   "Carrier_66_Motion_On_Fault" AT %Q3676.5 : Bool;
   "Carrier_66_Motion_Off_Fault" AT %Q3676.6 : Bool;
   "Carrier_66_Carrier_Spacing_Fault" AT %Q3676.7 : Bool;
   "Carrier_67_Carrier_In_Zone" AT %QW3700 : Word;
   "Carrier_67_Carrier_Number_Echo" AT %QW3702 : Word;
   "Carrier_67_Carrier_Position_Echo" AT %QD3704 : DWord;
   "Carrier_67_Next_Carrier_Number" AT %QW3708 : Word;
   "Carrier_67_Next_Stop_Position" AT %QD3710 : DWord;
   "Carrier_67_Drive_Command_Speed" AT %QW3714 : Word;
   "Carrier_67_Duplicate_Carrier_Number" AT %QW3716 : Word;
   "Carrier_67_First_Duplicate_Carrier_Position" AT %QD3718 : DWord;
   "Carrier_67_Second_Duplicate_Carrier_Position" AT %QD3722 : DWord;
   "Carrier_67_CommandWord" AT %QW3726 : Word;
   "Carrier_67_Heartbeat" AT %Q3726.0 : Bool;
   "Carrier_67_Drive_Forward_Command" AT %Q3726.1 : Bool;
   "Carrier_67_Fault_Reset" AT %Q3726.2 : Bool;
   "Carrier_67_At_Command_Position" AT %Q3726.3 : Bool;
   "Carrier_67_Duplicate_Carrier_Fault" AT %Q3726.4 : Bool;
   "Carrier_67_Motion_On_Fault" AT %Q3726.5 : Bool;
   "Carrier_67_Motion_Off_Fault" AT %Q3726.6 : Bool;
   "Carrier_67_Carrier_Spacing_Fault" AT %Q3726.7 : Bool;
   "Carrier_68_Carrier_In_Zone" AT %QW3750 : Word;
   "Carrier_68_Carrier_Number_Echo" AT %QW3752 : Word;
   "Carrier_68_Carrier_Position_Echo" AT %QD3754 : DWord;
   "Carrier_68_Next_Carrier_Number" AT %QW3758 : Word;
   "Carrier_68_Next_Stop_Position" AT %QD3760 : DWord;
   "Carrier_68_Drive_Command_Speed" AT %QW3764 : Word;
   "Carrier_68_Duplicate_Carrier_Number" AT %QW3766 : Word;
   "Carrier_68_First_Duplicate_Carrier_Position" AT %QD3768 : DWord;
   "Carrier_68_Second_Duplicate_Carrier_Position" AT %QD3772 : DWord;
   "Carrier_68_CommandWord" AT %QW3776 : Word;
   "Carrier_68_Heartbeat" AT %Q3776.0 : Bool;
   "Carrier_68_Drive_Forward_Command" AT %Q3776.1 : Bool;
   "Carrier_68_Fault_Reset" AT %Q3776.2 : Bool;
   "Carrier_68_At_Command_Position" AT %Q3776.3 : Bool;
   "Carrier_68_Duplicate_Carrier_Fault" AT %Q3776.4 : Bool;
   "Carrier_68_Motion_On_Fault" AT %Q3776.5 : Bool;
   "Carrier_68_Motion_Off_Fault" AT %Q3776.6 : Bool;
   "Carrier_68_Carrier_Spacing_Fault" AT %Q3776.7 : Bool;
   "Carrier_69_Carrier_In_Zone" AT %QW3800 : Word;
   "Carrier_69_Carrier_Number_Echo" AT %QW3802 : Word;
   "Carrier_69_Carrier_Position_Echo" AT %QD3804 : DWord;
   "Carrier_69_Next_Carrier_Number" AT %QW3808 : Word;
   "Carrier_69_Next_Stop_Position" AT %QD3810 : DWord;
   "Carrier_69_Drive_Command_Speed" AT %QW3814 : Word;
   "Carrier_69_Duplicate_Carrier_Number" AT %QW3816 : Word;
   "Carrier_69_First_Duplicate_Carrier_Position" AT %QD3818 : DWord;
   "Carrier_69_Second_Duplicate_Carrier_Position" AT %QD3822 : DWord;
   "Carrier_69_CommandWord" AT %QW3826 : Word;
   "Carrier_69_Heartbeat" AT %Q3826.0 : Bool;
   "Carrier_69_Drive_Forward_Command" AT %Q3826.1 : Bool;
   "Carrier_69_Fault_Reset" AT %Q3826.2 : Bool;
   "Carrier_69_At_Command_Position" AT %Q3826.3 : Bool;
   "Carrier_69_Duplicate_Carrier_Fault" AT %Q3826.4 : Bool;
   "Carrier_69_Motion_On_Fault" AT %Q3826.5 : Bool;
   "Carrier_69_Motion_Off_Fault" AT %Q3826.6 : Bool;
   "Carrier_69_Carrier_Spacing_Fault" AT %Q3826.7 : Bool;
   "Carrier_70_Carrier_In_Zone" AT %QW3850 : Word;
   "Carrier_70_Carrier_Number_Echo" AT %QW3852 : Word;
   "Carrier_70_Carrier_Position_Echo" AT %QD3854 : DWord;
   "Carrier_70_Next_Carrier_Number" AT %QW3858 : Word;
   "Carrier_70_Next_Stop_Position" AT %QD3860 : DWord;
   "Carrier_70_Drive_Command_Speed" AT %QW3864 : Word;
   "Carrier_70_Duplicate_Carrier_Number" AT %QW3866 : Word;
   "Carrier_70_First_Duplicate_Carrier_Position" AT %QD3868 : DWord;
   "Carrier_70_Second_Duplicate_Carrier_Position" AT %QD3872 : DWord;
   "Carrier_70_CommandWord" AT %QW3876 : Word;
   "Carrier_70_Heartbeat" AT %Q3876.0 : Bool;
   "Carrier_70_Drive_Forward_Command" AT %Q3876.1 : Bool;
   "Carrier_70_Fault_Reset" AT %Q3876.2 : Bool;
   "Carrier_70_At_Command_Position" AT %Q3876.3 : Bool;
   "Carrier_70_Duplicate_Carrier_Fault" AT %Q3876.4 : Bool;
   "Carrier_70_Motion_On_Fault" AT %Q3876.5 : Bool;
   "Carrier_70_Motion_Off_Fault" AT %Q3876.6 : Bool;
   "Carrier_70_Carrier_Spacing_Fault" AT %Q3876.7 : Bool;
   "Carrier_71_Carrier_In_Zone" AT %QW3900 : Word;
   "Carrier_71_Carrier_Number_Echo" AT %QW3902 : Word;
   "Carrier_71_Carrier_Position_Echo" AT %QD3904 : DWord;
   "Carrier_71_Next_Carrier_Number" AT %QW3908 : Word;
   "Carrier_71_Next_Stop_Position" AT %QD3910 : DWord;
   "Carrier_71_Drive_Command_Speed" AT %QW3914 : Word;
   "Carrier_71_Duplicate_Carrier_Number" AT %QW3916 : Word;
   "Carrier_71_First_Duplicate_Carrier_Position" AT %QD3918 : DWord;
   "Carrier_71_Second_Duplicate_Carrier_Position" AT %QD3922 : DWord;
   "Carrier_71_CommandWord" AT %QW3926 : Word;
   "Carrier_71_Heartbeat" AT %Q3926.0 : Bool;
   "Carrier_71_Drive_Forward_Command" AT %Q3926.1 : Bool;
   "Carrier_71_Fault_Reset" AT %Q3926.2 : Bool;
   "Carrier_71_At_Command_Position" AT %Q3926.3 : Bool;
   "Carrier_71_Duplicate_Carrier_Fault" AT %Q3926.4 : Bool;
   "Carrier_71_Motion_On_Fault" AT %Q3926.5 : Bool;
   "Carrier_71_Motion_Off_Fault" AT %Q3926.6 : Bool;
   "Carrier_71_Carrier_Spacing_Fault" AT %Q3926.7 : Bool;
   "Carrier_72_Carrier_In_Zone" AT %QW3950 : Word;
   "Carrier_72_Carrier_Number_Echo" AT %QW3952 : Word;
   "Carrier_72_Carrier_Position_Echo" AT %QD3954 : DWord;
   "Carrier_72_Next_Carrier_Number" AT %QW3958 : Word;
   "Carrier_72_Next_Stop_Position" AT %QD3960 : DWord;
   "Carrier_72_Drive_Command_Speed" AT %QW3964 : Word;
   "Carrier_72_Duplicate_Carrier_Number" AT %QW3966 : Word;
   "Carrier_72_First_Duplicate_Carrier_Position" AT %QD3968 : DWord;
   "Carrier_72_Second_Duplicate_Carrier_Position" AT %QD3972 : DWord;
   "Carrier_72_CommandWord" AT %QW3976 : Word;
   "Carrier_72_Heartbeat" AT %Q3976.0 : Bool;
   "Carrier_72_Drive_Forward_Command" AT %Q3976.1 : Bool;
   "Carrier_72_Fault_Reset" AT %Q3976.2 : Bool;
   "Carrier_72_At_Command_Position" AT %Q3976.3 : Bool;
   "Carrier_72_Duplicate_Carrier_Fault" AT %Q3976.4 : Bool;
   "Carrier_72_Motion_On_Fault" AT %Q3976.5 : Bool;
   "Carrier_72_Motion_Off_Fault" AT %Q3976.6 : Bool;
   "Carrier_72_Carrier_Spacing_Fault" AT %Q3976.7 : Bool;
   "Carrier_73_Carrier_In_Zone" AT %QW4000 : Word;
   "Carrier_73_Carrier_Number_Echo" AT %QW4002 : Word;
   "Carrier_73_Carrier_Position_Echo" AT %QD4004 : DWord;
   "Carrier_73_Next_Carrier_Number" AT %QW4008 : Word;
   "Carrier_73_Next_Stop_Position" AT %QD4010 : DWord;
   "Carrier_73_Drive_Command_Speed" AT %QW4014 : Word;
   "Carrier_73_Duplicate_Carrier_Number" AT %QW4016 : Word;
   "Carrier_73_First_Duplicate_Carrier_Position" AT %QD4018 : DWord;
   "Carrier_73_Second_Duplicate_Carrier_Position" AT %QD4022 : DWord;
   "Carrier_73_CommandWord" AT %QW4026 : Word;
   "Carrier_73_Heartbeat" AT %Q4026.0 : Bool;
   "Carrier_73_Drive_Forward_Command" AT %Q4026.1 : Bool;
   "Carrier_73_Fault_Reset" AT %Q4026.2 : Bool;
   "Carrier_73_At_Command_Position" AT %Q4026.3 : Bool;
   "Carrier_73_Duplicate_Carrier_Fault" AT %Q4026.4 : Bool;
   "Carrier_73_Motion_On_Fault" AT %Q4026.5 : Bool;
   "Carrier_73_Motion_Off_Fault" AT %Q4026.6 : Bool;
   "Carrier_73_Carrier_Spacing_Fault" AT %Q4026.7 : Bool;
   "Carrier_74_Carrier_In_Zone" AT %QW4050 : Word;
   "Carrier_74_Carrier_Number_Echo" AT %QW4052 : Word;
   "Carrier_74_Carrier_Position_Echo" AT %QD4054 : DWord;
   "Carrier_74_Next_Carrier_Number" AT %QW4058 : Word;
   "Carrier_74_Next_Stop_Position" AT %QD4060 : DWord;
   "Carrier_74_Drive_Command_Speed" AT %QW4064 : Word;
   "Carrier_74_Duplicate_Carrier_Number" AT %QW4066 : Word;
   "Carrier_74_First_Duplicate_Carrier_Position" AT %QD4068 : DWord;
   "Carrier_74_Second_Duplicate_Carrier_Position" AT %QD4072 : DWord;
   "Carrier_74_CommandWord" AT %QW4076 : Word;
   "Carrier_74_Heartbeat" AT %Q4076.0 : Bool;
   "Carrier_74_Drive_Forward_Command" AT %Q4076.1 : Bool;
   "Carrier_74_Fault_Reset" AT %Q4076.2 : Bool;
   "Carrier_74_At_Command_Position" AT %Q4076.3 : Bool;
   "Carrier_74_Duplicate_Carrier_Fault" AT %Q4076.4 : Bool;
   "Carrier_74_Motion_On_Fault" AT %Q4076.5 : Bool;
   "Carrier_74_Motion_Off_Fault" AT %Q4076.6 : Bool;
   "Carrier_74_Carrier_Spacing_Fault" AT %Q4076.7 : Bool;
   "Carrier_75_Carrier_In_Zone" AT %QW4100 : Word;
   "Carrier_75_Carrier_Number_Echo" AT %QW4102 : Word;
   "Carrier_75_Carrier_Position_Echo" AT %QD4104 : DWord;
   "Carrier_75_Next_Carrier_Number" AT %QW4108 : Word;
   "Carrier_75_Next_Stop_Position" AT %QD4110 : DWord;
   "Carrier_75_Drive_Command_Speed" AT %QW4114 : Word;
   "Carrier_75_Duplicate_Carrier_Number" AT %QW4116 : Word;
   "Carrier_75_First_Duplicate_Carrier_Position" AT %QD4118 : DWord;
   "Carrier_75_Second_Duplicate_Carrier_Position" AT %QD4122 : DWord;
   "Carrier_75_CommandWord" AT %QW4126 : Word;
   "Carrier_75_Heartbeat" AT %Q4126.0 : Bool;
   "Carrier_75_Drive_Forward_Command" AT %Q4126.1 : Bool;
   "Carrier_75_Fault_Reset" AT %Q4126.2 : Bool;
   "Carrier_75_At_Command_Position" AT %Q4126.3 : Bool;
   "Carrier_75_Duplicate_Carrier_Fault" AT %Q4126.4 : Bool;
   "Carrier_75_Motion_On_Fault" AT %Q4126.5 : Bool;
   "Carrier_75_Motion_Off_Fault" AT %Q4126.6 : Bool;
   "Carrier_75_Carrier_Spacing_Fault" AT %Q4126.7 : Bool;
   "Carrier_76_Carrier_In_Zone" AT %QW4150 : Word;
   "Carrier_76_Carrier_Number_Echo" AT %QW4152 : Word;
   "Carrier_76_Carrier_Position_Echo" AT %QD4154 : DWord;
   "Carrier_76_Next_Carrier_Number" AT %QW4158 : Word;
   "Carrier_76_Next_Stop_Position" AT %QD4160 : DWord;
   "Carrier_76_Drive_Command_Speed" AT %QW4164 : Word;
   "Carrier_76_Duplicate_Carrier_Number" AT %QW4166 : Word;
   "Carrier_76_First_Duplicate_Carrier_Position" AT %QD4168 : DWord;
   "Carrier_76_Second_Duplicate_Carrier_Position" AT %QD4172 : DWord;
   "Carrier_76_CommandWord" AT %QW4176 : Word;
   "Carrier_76_Heartbeat" AT %Q4176.0 : Bool;
   "Carrier_76_Drive_Forward_Command" AT %Q4176.1 : Bool;
   "Carrier_76_Fault_Reset" AT %Q4176.2 : Bool;
   "Carrier_76_At_Command_Position" AT %Q4176.3 : Bool;
   "Carrier_76_Duplicate_Carrier_Fault" AT %Q4176.4 : Bool;
   "Carrier_76_Motion_On_Fault" AT %Q4176.5 : Bool;
   "Carrier_76_Motion_Off_Fault" AT %Q4176.6 : Bool;
   "Carrier_76_Carrier_Spacing_Fault" AT %Q4176.7 : Bool;
   "Carrier_77_Carrier_In_Zone" AT %QW4200 : Word;
   "Carrier_77_Carrier_Number_Echo" AT %QW4202 : Word;
   "Carrier_77_Carrier_Position_Echo" AT %QD4204 : DWord;
   "Carrier_77_Next_Carrier_Number" AT %QW4208 : Word;
   "Carrier_77_Next_Stop_Position" AT %QD4210 : DWord;
   "Carrier_77_Drive_Command_Speed" AT %QW4214 : Word;
   "Carrier_77_Duplicate_Carrier_Number" AT %QW4216 : Word;
   "Carrier_77_First_Duplicate_Carrier_Position" AT %QD4218 : DWord;
   "Carrier_77_Second_Duplicate_Carrier_Position" AT %QD4222 : DWord;
   "Carrier_77_CommandWord" AT %QW4226 : Word;
   "Carrier_77_Heartbeat" AT %Q4226.0 : Bool;
   "Carrier_77_Drive_Forward_Command" AT %Q4226.1 : Bool;
   "Carrier_77_Fault_Reset" AT %Q4226.2 : Bool;
   "Carrier_77_At_Command_Position" AT %Q4226.3 : Bool;
   "Carrier_77_Duplicate_Carrier_Fault" AT %Q4226.4 : Bool;
   "Carrier_77_Motion_On_Fault" AT %Q4226.5 : Bool;
   "Carrier_77_Motion_Off_Fault" AT %Q4226.6 : Bool;
   "Carrier_77_Carrier_Spacing_Fault" AT %Q4226.7 : Bool;
   "Carrier_78_Carrier_In_Zone" AT %QW4250 : Word;
   "Carrier_78_Carrier_Number_Echo" AT %QW4252 : Word;
   "Carrier_78_Carrier_Position_Echo" AT %QD4254 : DWord;
   "Carrier_78_Next_Carrier_Number" AT %QW4258 : Word;
   "Carrier_78_Next_Stop_Position" AT %QD4260 : DWord;
   "Carrier_78_Drive_Command_Speed" AT %QW4264 : Word;
   "Carrier_78_Duplicate_Carrier_Number" AT %QW4266 : Word;
   "Carrier_78_First_Duplicate_Carrier_Position" AT %QD4268 : DWord;
   "Carrier_78_Second_Duplicate_Carrier_Position" AT %QD4272 : DWord;
   "Carrier_78_CommandWord" AT %QW4276 : Word;
   "Carrier_78_Heartbeat" AT %Q4276.0 : Bool;
   "Carrier_78_Drive_Forward_Command" AT %Q4276.1 : Bool;
   "Carrier_78_Fault_Reset" AT %Q4276.2 : Bool;
   "Carrier_78_At_Command_Position" AT %Q4276.3 : Bool;
   "Carrier_78_Duplicate_Carrier_Fault" AT %Q4276.4 : Bool;
   "Carrier_78_Motion_On_Fault" AT %Q4276.5 : Bool;
   "Carrier_78_Motion_Off_Fault" AT %Q4276.6 : Bool;
   "Carrier_78_Carrier_Spacing_Fault" AT %Q4276.7 : Bool;
   "Carrier_79_Carrier_In_Zone" AT %QW4300 : Word;
   "Carrier_79_Carrier_Number_Echo" AT %QW4302 : Word;
   "Carrier_79_Carrier_Position_Echo" AT %QD4304 : DWord;
   "Carrier_79_Next_Carrier_Number" AT %QW4308 : Word;
   "Carrier_79_Next_Stop_Position" AT %QD4310 : DWord;
   "Carrier_79_Drive_Command_Speed" AT %QW4314 : Word;
   "Carrier_79_Duplicate_Carrier_Number" AT %QW4316 : Word;
   "Carrier_79_First_Duplicate_Carrier_Position" AT %QD4318 : DWord;
   "Carrier_79_Second_Duplicate_Carrier_Position" AT %QD4322 : DWord;
   "Carrier_79_CommandWord" AT %QW4326 : Word;
   "Carrier_79_Heartbeat" AT %Q4326.0 : Bool;
   "Carrier_79_Drive_Forward_Command" AT %Q4326.1 : Bool;
   "Carrier_79_Fault_Reset" AT %Q4326.2 : Bool;
   "Carrier_79_At_Command_Position" AT %Q4326.3 : Bool;
   "Carrier_79_Duplicate_Carrier_Fault" AT %Q4326.4 : Bool;
   "Carrier_79_Motion_On_Fault" AT %Q4326.5 : Bool;
   "Carrier_79_Motion_Off_Fault" AT %Q4326.6 : Bool;
   "Carrier_79_Carrier_Spacing_Fault" AT %Q4326.7 : Bool;
   "Carrier_80_Carrier_In_Zone" AT %QW4350 : Word;
   "Carrier_80_Carrier_Number_Echo" AT %QW4352 : Word;
   "Carrier_80_Carrier_Position_Echo" AT %QD4354 : DWord;
   "Carrier_80_Next_Carrier_Number" AT %QW4358 : Word;
   "Carrier_80_Next_Stop_Position" AT %QD4360 : DWord;
   "Carrier_80_Drive_Command_Speed" AT %QW4364 : Word;
   "Carrier_80_Duplicate_Carrier_Number" AT %QW4366 : Word;
   "Carrier_80_First_Duplicate_Carrier_Position" AT %QD4368 : DWord;
   "Carrier_80_Second_Duplicate_Carrier_Position" AT %QD4372 : DWord;
   "Carrier_80_CommandWord" AT %QW4376 : Word;
   "Carrier_80_Heartbeat" AT %Q4376.0 : Bool;
   "Carrier_80_Drive_Forward_Command" AT %Q4376.1 : Bool;
   "Carrier_80_Fault_Reset" AT %Q4376.2 : Bool;
   "Carrier_80_At_Command_Position" AT %Q4376.3 : Bool;
   "Carrier_80_Duplicate_Carrier_Fault" AT %Q4376.4 : Bool;
   "Carrier_80_Motion_On_Fault" AT %Q4376.5 : Bool;
   "Carrier_80_Motion_Off_Fault" AT %Q4376.6 : Bool;
   "Carrier_80_Carrier_Spacing_Fault" AT %Q4376.7 : Bool;
   "Carrier_81_Carrier_In_Zone" AT %QW4400 : Word;
   "Carrier_81_Carrier_Number_Echo" AT %QW4402 : Word;
   "Carrier_81_Carrier_Position_Echo" AT %QD4404 : DWord;
   "Carrier_81_Next_Carrier_Number" AT %QW4408 : Word;
   "Carrier_81_Next_Stop_Position" AT %QD4410 : DWord;
   "Carrier_81_Drive_Command_Speed" AT %QW4414 : Word;
   "Carrier_81_Duplicate_Carrier_Number" AT %QW4416 : Word;
   "Carrier_81_First_Duplicate_Carrier_Position" AT %QD4418 : DWord;
   "Carrier_81_Second_Duplicate_Carrier_Position" AT %QD4422 : DWord;
   "Carrier_81_CommandWord" AT %QW4426 : Word;
   "Carrier_81_Heartbeat" AT %Q4426.0 : Bool;
   "Carrier_81_Drive_Forward_Command" AT %Q4426.1 : Bool;
   "Carrier_81_Fault_Reset" AT %Q4426.2 : Bool;
   "Carrier_81_At_Command_Position" AT %Q4426.3 : Bool;
   "Carrier_81_Duplicate_Carrier_Fault" AT %Q4426.4 : Bool;
   "Carrier_81_Motion_On_Fault" AT %Q4426.5 : Bool;
   "Carrier_81_Motion_Off_Fault" AT %Q4426.6 : Bool;
   "Carrier_81_Carrier_Spacing_Fault" AT %Q4426.7 : Bool;
   "Carrier_82_Carrier_In_Zone" AT %QW4450 : Word;
   "Carrier_82_Carrier_Number_Echo" AT %QW4452 : Word;
   "Carrier_82_Carrier_Position_Echo" AT %QD4454 : DWord;
   "Carrier_82_Next_Carrier_Number" AT %QW4458 : Word;
   "Carrier_82_Next_Stop_Position" AT %QD4460 : DWord;
   "Carrier_82_Drive_Command_Speed" AT %QW4464 : Word;
   "Carrier_82_Duplicate_Carrier_Number" AT %QW4466 : Word;
   "Carrier_82_First_Duplicate_Carrier_Position" AT %QD4468 : DWord;
   "Carrier_82_Second_Duplicate_Carrier_Position" AT %QD4472 : DWord;
   "Carrier_82_CommandWord" AT %QW4476 : Word;
   "Carrier_82_Heartbeat" AT %Q4476.0 : Bool;
   "Carrier_82_Drive_Forward_Command" AT %Q4476.1 : Bool;
   "Carrier_82_Fault_Reset" AT %Q4476.2 : Bool;
   "Carrier_82_At_Command_Position" AT %Q4476.3 : Bool;
   "Carrier_82_Duplicate_Carrier_Fault" AT %Q4476.4 : Bool;
   "Carrier_82_Motion_On_Fault" AT %Q4476.5 : Bool;
   "Carrier_82_Motion_Off_Fault" AT %Q4476.6 : Bool;
   "Carrier_82_Carrier_Spacing_Fault" AT %Q4476.7 : Bool;
END_VAR

TYPE "UDT_SDCOutFaults"
VERSION : 0.1
   STRUCT
      DuplicateCarrierFault : Bool;
      MotionOnFault : Bool;
      MotionOffFault : Bool;
      CarrierSpacingFault : Bool;
   END_STRUCT;
END_TYPE

TYPE "UDT_Stop"
VERSION : 0.1
   STRUCT
      StopNumber : Bool;
      StopPosition : Bool;
      ClearToRelease : Bool;
      CarrierPresentStop : Bool;
   END_STRUCT;
END_TYPE

TYPE "UDT_HMIZonePositionStructure"
   STRUCT
      ZonePosition : Word;
      CarrierNumber : Word;
      CarrierPosition : Word;
      Faulted : Bool;
   END_STRUCT;
END_TYPE

TYPE "UDT_System"
VERSION : 0.1
   STRUCT
      Zone : Array[0..65] of "UDT_ZoneStructure";
      Carrier : Array[0..99] of "UDT_CarrierStructure";
      LowSpeedSetpoint : Word;
      HighSpeedSetpoint : Word;
      DecelPositionOffset : Word;
      SDC_Faults : Array[0..9] of Int;
      Carrier_Spacing : Int;
      TotalZones : Int;
      TotalZonePosn : Int;
      TotalCarriers : Int;
      CoarsePositionTolerance : Word;
      FinePositionTolerance : Word;
      CoarsePositionDecelOffset : Word;
      FinePositionDecelOffset : Word;
      Production_Spacing : Word;
      ClearOfStopDist : Word;
      FineDecelSpeed : Word;
      CoarseDecelSpeed : Word;
      ProductionZnSpeed : Word;
      AccumZnSpeed : Word;
      SDC : "UDT_SDC";
   END_STRUCT;
END_TYPE

TYPE "UDT_Carrier"
VERSION : 0.1
   STRUCT
      CARRIER : Array[1..99] of "UDT_CarrierStructure";
   END_STRUCT;
END_TYPE

TYPE "UDT_SDC_IN"
VERSION : 0.1
   STRUCT
      CarrierNumber : Word;
      CarrierPosition : DWord;
      ActualSpeed : Word;
      CarrierDriveFaults : Word;
      CarrierDriveAlarms : Word;
      CarrierFaults : Word;
      Spare_Word : Word;
      RunningFWD : Bool;
      RunningREV : Bool;
      Stopped : Bool;
      ProductionHoldPB_Status : Bool;
      CrashDetectStatus : Bool;
      HeartBeat : Bool;
      AutoMode : Bool;
      ManualMode : Bool;
      IR_Remote_9_Pressed : Bool;
      EncoderCommFault : Bool;
      DriveCommFault : Bool;
      HMICommFault : Bool;
   END_STRUCT;
END_TYPE

TYPE "UDT_SDC_OUT"
VERSION : 0.1
   STRUCT
      Zone : Int;
      CarrierNum : Word;
      CarrierPosition : DWord;
      NextCarrierNum : Word;
      NextStopPos : DWord;
      DriveFwdCMD : Bool;
      DriveCmdSpeed : Word;
      Spare_Word_1 : Word;
      Spare_Word_2 : Word;
      HeartBeat : Bool;
      FaultReset : Bool;
      HighSpeedEnable : Bool;
      AtCmdPos : Bool;
      DuplicateCarrierNum : Word;
      FirstDuplicateFndPos : Bool;
      SecondDuplicateFndPos : Bool;
      Faults : "UDT_SDCOutFaults";
   END_STRUCT;
END_TYPE

TYPE "UDT_CarrierFaults"
VERSION : 0.1
   STRUCT
      Fault : Array[0..9] of Int;
   END_STRUCT;
END_TYPE

TYPE "UDT_SDC"
   STRUCT
      HMI : "UDT_Drive_HMI";
   END_STRUCT;
END_TYPE

TYPE "UDT_TrafficCop"
VERSION : 0.1
   STRUCT
      Element_1 : Bool;
      AutoSpeedFast : Word;
      AutoSpeedSlow : Word;
      CommandPosLowLimit : DWord;
      CommandPosHighLimit : DWord;
      CommandPos : DWord;
      AtCommandPos : Bool;
      DecelPosition : DWord;
   END_STRUCT;
END_TYPE

TYPE "UDT_SDC_6EMS_TS_STAT"
VERSION : 0.1
   STRUCT
      EMS : Array[1..6] of "UDT_SDC_EMS_TS_STAT";
   END_STRUCT;
END_TYPE

TYPE "UDT_SDC_6EMS_TS_STAT_HMI"
VERSION : 0.1
   STRUCT
      EMS : Array[1..6] of "UDT_SDC_EMS_TS_STAT_HMI";
   END_STRUCT;
END_TYPE

TYPE "UDT_EMS_IF_Q_VFC"
VERSION : 0.1
   STRUCT
      VFC_No : Byte;   // FU Nummer (z.B.: 1=Fahren, 2=Heben, 3=Schwenken) / VFC number (f.e.: 1=Drive, 2=Hoist, 3=Tilt)
      PW1 : Word;   // Prozesswort 1 / Processdataword 1
      PW2 : Word;   // Prozesswort 2 / Processdataword 2
      PW3 : Word;   // Prozesswort 3 / Processdataword 3
   END_STRUCT;
END_TYPE

TYPE "UDT_EMS_TA"
VERSION : 0.1
   STRUCT
      ZSW1 : Word;   // G120D Zustandswort 1 / Statusword 1
      ERROR : Word;   // G120D Störcode / Errorcode
      CURRENT : Word;   // G120D Strom / Current
      FAULT : Word;   // G120D Störcode / Errorcode
      ALARM : Word;
   END_STRUCT;
END_TYPE

TYPE "UDT_EMS_IF_Q_IQ"
VERSION : 0.1
   STRUCT
      BS1PH1_KANAL_1 : Bool;
      BS1PH1_KANAL_2 : Bool;
      BS1PH1_KANAL_3 : Bool;
      BS1PH1_KANAL_4 : Bool;
      BS1PH1_KANAL_5 : Bool;
      BS1PH1_KANAL_6 : Bool;
      BS1PH1_KANAL_7 : Bool;
      BS1PH1_KANAL_8 : Bool;
      BS1FC302 : Bool;
      AB1FCM1 : Bool;
      AB1QA1_R : Bool;
      I_1_3 : Bool;
      I_1_8 : Bool;
      I_1_5 : Bool;
      I_1_6 : Bool;
      I_1_7 : Bool;
      HE1BGS03a : Bool;
      HE1BGS03b : Bool;
      HE1BGS05 : Bool;
      BS1SFWE2 : Bool;
      I_2_4 : Bool;
      I_2_5 : Bool;
      I_2_6 : Bool;
      I_2_7 : Bool;
      I_6_0 : Bool;
      I_6_1 : Bool;
      I_6_2 : Bool;
      I_6_3 : Bool;
      I_6_4 : Bool;
      I_6_5 : Bool;
      I_6_6 : Bool;
      I_6_7 : Bool;
      "BS1PH1_L+" : Bool;
      BS1PH1_DAT : Bool;
      AB1QA1 : Bool;
      O_0_3 : Bool;
      O_0_4 : Bool;
      O_0_5 : Bool;
      O_0_6 : Bool;
      O_0_7 : Bool;
      HE1KK1 : Bool;
      O_8_1 : Bool;
      O_8_2 : Bool;
      O_8_3 : Bool;
      O_8_4 : Bool;
      O_8_5 : Bool;
      O_8_6 : Bool;
      O_8_7 : Bool;
      I_261_0 : Bool;
      I_261_1 : Bool;
      I_261_2 : Bool;
      I_261_3 : Bool;
      I_261_4 : Bool;
      I_261_5 : Bool;
      I_261_6 : Bool;
      I_261_7 : Bool;
      HE1BGG1 : Bool;
      "HE1BGG1:13" : Bool;
      HE1BGE05 : Bool;
      I_271_3 : Bool;
      I_271_4 : Bool;
      I_271_5 : Bool;
      I_271_6 : Bool;
      I_271_7 : Bool;
      SN1BGE04 : Bool;
      I_281_1 : Bool;
      I_281_2 : Bool;
      I_281_3 : Bool;
      I_281_4 : Bool;
      I_281_5 : Bool;
      I_281_6 : Bool;
      I_281_7 : Bool;
      I_285_0 : Bool;
      I_285_1 : Bool;
      I_285_2 : Bool;
      I_285_3 : Bool;
      I_285_4 : Bool;
      I_285_5 : Bool;
      I_285_6 : Bool;
      I_285_7 : Bool;
   END_STRUCT;
END_TYPE

TYPE "UDT_SDC_EMS_TS_STAT_HMI"
VERSION : 0.1
   STRUCT
      EMS_ID : Int;
      PROFILE : Int;
      DRIVE_POS : DInt;
      HOIST_POS : Int;
      ERROR : Int;
      "DRIVE_POS_%" : Int;
      SEK_NR : Int;
      STAT_1 : DWord;
      STAT_2 : Word;
      SORTE : DWord;
      FKT : DWord;
   END_STRUCT;
END_TYPE

TYPE "UDT_SDC_FT_STAT"
VERSION : 0.1
   STRUCT
      STAT : Array[1..4] of "UDT_SDC_EMS_TS_STAT";
   END_STRUCT;
END_TYPE

TYPE "UDT_EMS_IF_I"
VERSION : 0.1
   STRUCT
      EMS_ID : Int;   // EMS Nummer / EMS number
      CONT : "UDT_EMS_IF_I_CONTR";   // Steuerbit`s / Controlbit`s
      D_SETPOS : DInt;   // Sollposition Fahrantrieb / setpoint drive position (mm)
      D_SETSPEED : DInt;   // Sollgeschwindigkeit Fahrantrieb / set value drive speed (mm/min)
      H_SETPOS : Int;   // Sollposition Hubantrieb / setpoint hoist position (mm)
      H_SETSPEED : Int;   // Sollgeschwindigkeit Hubantrieb / setpoint hoist speed (mm/min)
      Reserve18 : Int;
      Reserve20 : Int;
      FB_VFC_No : Byte;   // Rückmeldung Prozesswerte FU`s / Feedback VFC PDAT
      FB_ER_WORD_No : Int;   // Rückmeldung Zähler Störnummern / Feedback Transfer counter error words
      DB_No : Int;   // DB Nummer Datentransfer / DB No. data transfer
      DBB_No : Int;   // DBB Nummer Datentransfer / DBB No. data transfer
      DB_UserData : DWord;   // Nutzdaten Datentransfer / User data, data transfer
      ERRORS_SPLC : "UDT_EMS_IF_I_SDC_ERRORS";   // Störungen Kopfsteuerung / Errors from System-PLC
      Reserve36 : Word;   // Reserve / spare
      Reserve38 : Word;   // Reserve / spare
   END_STRUCT;
END_TYPE

TYPE "UDT_EMS_PAR"
VERSION : 0.1
   STRUCT
      DRIVE : Struct
         Funct : Struct   // several functions
            Res0 : Bool := TRUE;   // Reserve: without swich-off Scanner
            IgnoreBridgeStopp : Bool := TRUE;   // Ignore Bridge Stopp-Position after Startpoint for Positioning
            DontIgnoreAPOSwhenDriving : Bool := FALSE;   // spare
            Speed0_1mm_s : Bool := FALSE;   // spare
            IR_noEMSnumber : Bool := FALSE;   // spare
            IR_noLogin : Bool := FALSE;   // spare
            Res6 : Bool := FALSE;   // spare
            Res7 : Bool := FALSE;   // spare
            Res8 : Bool := FALSE;   // spare
            Res9 : Bool := FALSE;   // spare
            Res10 : Bool := FALSE;   // spare
            Res11 : Bool := FALSE;   // spare
            Res12 : Bool := FALSE;   // spare
            Res13 : Bool := FALSE;   // spare
            Res14 : Bool := FALSE;   // spare
            Res15 : Bool := FALSE;   // spare
         END_STRUCT;
         V_FACT_1 : Real := 0.00266;
         V_SETP_1 : DInt := 600;   // Setpoint for calculation of factor
         V_FACT_2 : Real := 0.00246;
         V_SETP_2 : DInt := 3000;   // Setpoint for calculation of factor
         V_FACT_3 : Real := 0.00246;
         V_SETP_3 : DInt := 10000;   // Setpoint for calculation of factor
         V_FACT_4 : Real := 0.00236;
         V_SETP_4 : DInt := 20000;   // Setpoint for calculation of factor
         V_LIMIT_FACT : Real := 0.3;
         V_FACT_5 : Real := 0.00226;
         "V_FACT_ACT_V_<600" : Real := 0.0027;   // Factor for conversion of mm/min to U/min -> determined
         "V_FACT_ACT_V_<1200" : Real := 0.0027;   // Factor for conversion of mm/min to U/min -> determined
         V_min : DInt := 500;   // minimum speed in mm/min
         V_max_top : DInt := 36000;   // maximum speed if hoist raised in mm/min
         V_max_Not_top : DInt := 16000;   // maximum speed if hoist not raised in mm/min
         V_Pos_1_Reserve : DInt := 0;   // Positioning speed 1 / Positioning with position setpoint
         V_Pos_2 : DInt := 10000;   // Positioning speed 2 / Positioning with position setpoint
         V_Pos_3_Reserve : DInt := 12000;   // Positioning speed 3 / Positioning with position setpoint
         V_Fixed_1 : DInt := 3000;   // Fixed speed 1 in mm/min (IR manual)
         V_Fixed_2 : DInt := 13000;   // Fixed speed 2 in mm/min (IR manual)
         V_Fixed_3_Reserve : DInt := 18000;   // Fixed speed 3 in mm/min
         V_Fixed_4_SLS_SPEED : DInt := 15000;   // Fixed speed 4 in mm/min V_SafeSpeed
         V_DIV_FAST : DInt := 18000;   // speed for Divisor positioning fast
         DIV_POS_FAST : DInt := 40;   // Divisor to calculate braking distance for positioning fast (>=18m/min)
         DIV_POS_SLOW : DInt := 60;   // Divisor to calculate braking distance for positioning slow (<18m/min)
         TOL_SET_POS : Int := 2;   // tolerance (mm) for setting the position signal
         TOL_RESET_POS : Int := 6;   // tolerance (mm) for resetting the position signal
         Window_Pos : Int := 2;   // Window (mm) for shut-down during positioning
         Window_Overrun : Int := 6;   // Window (mm) for check "Stop Position overrun"
         Window_Pos_2 : Int := 800;   // Window (mm) for switching to positioning speed 2
         Window_Movement : Int := 10;   // Window (mm) for check "Movement without release"
         Window_Distance_Reserve : Int := 10;   // Window (mm) for distance controller
         Delay_Pos : Int := 2000;   // Delay EMS in position (ms)
         Reserve_118 : S5Time := S5T#5M;   // Delay Barcode scanner off
         Reserve_120 : S5Time := S5T#2M;   // Delay Barcode scanner on
         DelaySpeedContr : S5Time := S5T#9S_900MS;   // Delay for speed control
         TolSpeedContr : Int := 60;   // tolerance for speed control (in %)
         SYNCH_MID_VALUE : Int := 60;   // spare
         SYNCH_tINCREASE : Int := 30;
      END_STRUCT;
      Reserve : Array[1..5] of Word;
      HOIST : Struct
         V_Min : Int := 200;   // minimum speed in mm/min
         V_Max : Int := 8000;   // maximum speed in mm/min
         V_MaxOccLift : Int := 6600;   // maximum speed in mm/min occupied lifitng
         V_Reserve_2 : Int := 0;   // hoist speed spare
         V_Pos_1 : Int := 800;   // Positioning speed1
         V_Pos_2 : Int := 2000;   // Positioning speed 2
         V_Fixed_1 : Int := 2000;   // Fixed speed 1 in mm/min (IR manual)
         V_Fixed_2 : Int := 4000;   // Fixed speed 2 in mm/min (IR manual)
         V_Fixed_3_START : Int := 200;   // Fixed speed 3 in mm/min
         V_Fixed_4_SLS_SPEED : Int := 2000;   // Fixed speed 4 in mm/min
         V_Fixed_5_Reserve : Int := 2000;   // slow safe speed (2000)
         V_Fixed_6_SlowSpeed : Int := 4000;   // Global Speed paramter for TS {"DB_SDC_COMMAND".Section[1].Commands.hoist_slow}
         V_FACT_Hz_UP : Real := 0.01246;   // Factor for conversion of current value from converter in % to mm/min
         V_FACT_Hz_DOWN : Real := 0.01246;   // Factor for conversion of current value from converter in % to mm/min
         H_Window_POS_V1 : Int := 20;   // Window (mm) for switching to positioning speed 1
         H_Window_POS_V2 : Int := 140;   // Window (mm) for switching to positioning speed 2
         H_TOL_SET_POS : Int := 2;   // tolerance (mm) for setting the position signal
         H_TOL_RESET_POS : Int := 8;   // tolerance (mm) for resetting the position signal
         H_MIN : Int := 4;   // minimum height
         H_MIN_without_bypass : Int := 126;   // minimum height without bypass switch (120)
         H_REF_OFFSET : Int := 9;   // Offset to hoist position reference prox.switch
         H_REF : Int := 2641;   // Height reference initiator Position
         H_FACT_ENC1 : Real := 1.0;   // Factor for conversion of encoder value in mm / encoder 1
         H_FACT_ENC2 : Real := 1.0;   // Factor for conversion of encoder value in mm / encoder 2
         H_FACT_SPEED : Real := 0.316;   // Factor for conversion of encoder value / encoder 1or2 in mm for speed
         H_ENC_MAX_DIFF : Int := 50;   // maximum difference between encoders
         H_Slow : Int := 660;   // slow height (500)
         H_tIN_POS : Int := 1000;   // Delay HOIST in position (ms)
         H_REF_HMI : Int := 2641;   // Height HMI reference
      END_STRUCT;
      Reserve1 : Array[1..6] of Word;
      TILT : Array[1..34] of Word;
      Reserve2 : Array[1..6] of Word;
   END_STRUCT;
   // Reserve1[6] := 16#0000;
   // Reserve1[5] := 16#0000;
   // Reserve1[4] := 16#0000;
   // Reserve1[3] := 16#0000;
   // Reserve1[2] := 16#0000;
   // Reserve1[1] := 16#0000;
   // Reserve[5] := 16#0000;
   // Reserve[4] := 16#0000;
   // Reserve[3] := 16#0000;
   // Reserve[2] := 16#0000;
   // Reserve[1] := 16#0000;
   // Reserve2[1] := 16#0000;
   // Reserve2[2] := 16#0000;
   // Reserve2[3] := 16#0000;
   // Reserve2[4] := 16#0000;
   // Reserve2[5] := 16#0000;
   // Reserve2[6] := 16#0000;
END_TYPE

TYPE "UDT_TrafficCopCarrierStructure"
VERSION : 0.1
   STRUCT
      MoveFwd : Bool;
      DriveCmdSpeed : Word;
      CommandPos : DWord;
      AtCmdPos : Bool;
      NextStopPos : DWord;
      NextCarrierNumber : Word;
      CarrierNumber : Word;
   END_STRUCT;
END_TYPE

TYPE "UDT_TrafficCopZoneStructure"
VERSION : 0.1
   STRUCT
      Carrier : Array[0..99] of "UDT_TrafficCopCarrierStructure";
   END_STRUCT;
END_TYPE

TYPE "UDT_SDC_FT_COM"
VERSION : 0.1
   STRUCT
      COM : Array[1..7] of "UDT_SDC_EMS_TS_COM";
   END_STRUCT;
END_TYPE

TYPE "UDT_TC_ZoneMotion"
VERSION : 0.1
   STRUCT
      Zone : Array[0..60] of "UDT_ZnPosMotion";
   END_STRUCT;
END_TYPE

TYPE "UDT_TC_ZnPosMotion"
VERSION : 0.1
   STRUCT
      zone : Array[0..60] of "UDT_TrafficCopZnPosStructure";
   END_STRUCT;
END_TYPE

TYPE "UDT_ZnPosMotion"
VERSION : 0.1
   STRUCT
      ZonePos : Array[0..99] of "UDT_TrafficCopCarrierStructure";
   END_STRUCT;
END_TYPE

TYPE "UDT_HMIZonePositions"
   STRUCT
      ZonePosition : Word;
   END_STRUCT;
END_TYPE

TYPE "UDT_TC_SDCOutZone"
VERSION : 0.1
   STRUCT
      Carrier : Array[0..99] of "UDT_TC_SDCOutCarrier";
   END_STRUCT;
END_TYPE

TYPE "UDT_Drive_HMI"
   STRUCT
      G120D_STATUS : Word;
      G120D_CONTROL : Word;
   END_STRUCT;
END_TYPE

TYPE "UDT_TC_SDC_Out"
VERSION : 0.1
   STRUCT
      Zone : Array[0..60] of "UDT_TC_SDCOutZone";
   END_STRUCT;
END_TYPE

TYPE "UDT_TC_SDCOutCarrier"
VERSION : 0.1
   STRUCT
      DriveFwdCMD : Bool;
      DriveCmdSpeed : Int;
      NextStopPos : DWord;
      NextCarrierNum : Word;
      AtCmdPos : Bool;
   END_STRUCT;
END_TYPE

TYPE "UDT_IN"
   STRUCT
      G120D_CONTROL : "UDT_G120D_ZSW1_STATUS";
      G120D_STATUS : "UDT_G120D_STW1_CONTROL";
      DecrementCarrierIndex : Bool;
      IncrementCarrierIndex : Bool;
      CarrierStatusIndex : Int;
      DecrementStatusIndex : Bool;
      IncrementStatusIndex : Bool;
      DriveStatusIndex : Int;
      DecrementZoneIndex : Bool;
      IncrementZoneIndex : Bool;
      ZoneStatusIndex : Int;
   END_STRUCT;
END_TYPE

TYPE "UDT_TrafficCopZnPosStructure"
VERSION : 0.1
   STRUCT
      ZonePos : Array[0..40] of "UDT_TrafficCopZoneStructure";
   END_STRUCT;
END_TYPE

